(* Logix 5000 project; controller UOWHF Emulate 5570 rev 30.12; software revision 30.00 *) (continued)
   		UOWHF_Add_c.2:=UOWHF_Result[2].31;
   		UOWHF_Result[2].31:=0;
   		UOWHF_Result[3]:=UOWHF_Result[3] + 1798644847+UOWHF_Add_c;
   		UOWHF_Add_c.3:=UOWHF_Result[3].31;
   		UOWHF_Result[3].31:=0;
   		UOWHF_Result[4]:=UOWHF_Result[4] + 304175449+UOWHF_Add_c;
   		UOWHF_Add_c.4:=UOWHF_Result[4].31;
   		UOWHF_Result[4].31:=0;
   	End_If;
   	If UOWHF_Msg[2].[30] Then
   		UOWHF_Result[0]:=UOWHF_Result[0] + 1161935431+UOWHF_Add_c;
   		UOWHF_Add_c.0:=UOWHF_Result[0].31;
   		UOWHF_Result[0].31:=0;
   		UOWHF_Result[1]:=UOWHF_Result[1] + 944693816+UOWHF_Add_c;
   		UOWHF_Add_c.1:=UOWHF_Result[1].31;
   		UOWHF_Result[1].31:=0;
   		UOWHF_Result[2]:=UOWHF_Result[2] + 1100985340+UOWHF_Add_c;
   		UOWHF_Add_c.2:=UOWHF_Result[2].31;
   		UOWHF_Result[2].31:=0;
   		UOWHF_Result[3]:=UOWHF_Result[3] + 216963659+UOWHF_Add_c;
   		UOWHF_Add_c.3:=UOWHF_Result[3].31;
   		UOWHF_Result[3].31:=0;
   		UOWHF_Result[4]:=UOWHF_Result[4] + 89876541+UOWHF_Add_c;
   		UOWHF_Add_c.4:=UOWHF_Result[4].31;
   		UOWHF_Result[4].31:=0;
   	End_If;
   	If UOWHF_Msg[2].[31] Then
   		UOWHF_Result[0]:=UOWHF_Result[0] + 1158699558+UOWHF_Add_c;
   		UOWHF_Add_c.0:=UOWHF_Result[0].31;
   		UOWHF_Result[0].31:=0;
   		UOWHF_Result[1]:=UOWHF_Result[1] + 148835756+UOWHF_Add_c;
   		UOWHF_Add_c.1:=UOWHF_Result[1].31;
   		UOWHF_Result[1].31:=0;
   		UOWHF_Result[2]:=UOWHF_Result[2] + 32681667+UOWHF_Add_c;
   		UOWHF_Add_c.2:=UOWHF_Result[2].31;
   		UOWHF_Result[2].31:=0;
   		UOWHF_Result[3]:=UOWHF_Result[3] + 636137273+UOWHF_Add_c;
   		UOWHF_Add_c.3:=UOWHF_Result[3].31;
   		UOWHF_Result[3].31:=0;
   		UOWHF_Result[4]:=UOWHF_Result[4] + 1474642829+UOWHF_Add_c;
   		UOWHF_Add_c.4:=UOWHF_Result[4].31;
   		UOWHF_Result[4].31:=0;
   	End_If;
   	If UOWHF_Msg[3].[0] Then
   		UOWHF_Result[0]:=UOWHF_Result[0] + 1085349533+UOWHF_Add_c;
   		UOWHF_Add_c.0:=UOWHF_Result[0].31;
   		UOWHF_Result[0].31:=0;
   		UOWHF_Result[1]:=UOWHF_Result[1] + 1302835678+UOWHF_Add_c;
   		UOWHF_Add_c.1:=UOWHF_Result[1].31;
   		UOWHF_Result[1].31:=0;
   		UOWHF_Result[2]:=UOWHF_Result[2] + 681913251+UOWHF_Add_c;
   		UOWHF_Add_c.2:=UOWHF_Result[2].31;
   		UOWHF_Result[2].31:=0;
   		UOWHF_Result[3]:=UOWHF_Result[3] + 723730247+UOWHF_Add_c;
   		UOWHF_Add_c.3:=UOWHF_Result[3].31;
   		UOWHF_Result[3].31:=0;
   		UOWHF_Result[4]:=UOWHF_Result[4] + 7919506+UOWHF_Add_c;
   		UOWHF_Add_c.4:=UOWHF_Result[4].31;
   		UOWHF_Result[4].31:=0;
   	End_If;
   	If UOWHF_Msg[3].[1] Then
   		UOWHF_Result[0]:=UOWHF_Result[0] + 1136561897+UOWHF_Add_c;
   		UOWHF_Add_c.0:=UOWHF_Result[0].31;
   		UOWHF_Result[0].31:=0;
   		UOWHF_Result[1]:=UOWHF_Result[1] + 1822763236+UOWHF_Add_c;
   		UOWHF_Add_c.1:=UOWHF_Result[1].31;
   		UOWHF_Result[1].31:=0;
   		UOWHF_Result[2]:=UOWHF_Result[2] + 2116802572+UOWHF_Add_c;
   		UOWHF_Add_c.2:=UOWHF_Result[2].31;
   		UOWHF_Result[2].31:=0;
   		UOWHF_Result[3]:=UOWHF_Result[3] + 595130731+UOWHF_Add_c;
   		UOWHF_Add_c.3:=UOWHF_Result[3].31;
   		UOWHF_Result[3].31:=0;
   		UOWHF_Result[4]:=UOWHF_Result[4] + 1143215041+UOWHF_Add_c;
   		UOWHF_Add_c.4:=UOWHF_Result[4].31;
   		UOWHF_Result[4].31:=0;
   	End_If;
   	If UOWHF_Msg[3].[2] Then
   		UOWHF_Result[0]:=UOWHF_Result[0] + 44711483+UOWHF_Add_c;
   		UOWHF_Add_c.0:=UOWHF_Result[0].31;
   		UOWHF_Result[0].31:=0;
   		UOWHF_Result[1]:=UOWHF_Result[1] + 757400375+UOWHF_Add_c;
   		UOWHF_Add_c.1:=UOWHF_Result[1].31;
   		UOWHF_Result[1].31:=0;
   		UOWHF_Result[2]:=UOWHF_Result[2] + 1986965253+UOWHF_Add_c;
   		UOWHF_Add_c.2:=UOWHF_Result[2].31;
   		UOWHF_Result[2].31:=0;
   		UOWHF_Result[3]:=UOWHF_Result[3] + 1261883823+UOWHF_Add_c;
   		UOWHF_Add_c.3:=UOWHF_Result[3].31;
   		UOWHF_Result[3].31:=0;
   		UOWHF_Result[4]:=UOWHF_Result[4] + 1629162798+UOWHF_Add_c;
   		UOWHF_Add_c.4:=UOWHF_Result[4].31;
   		UOWHF_Result[4].31:=0;
   	End_If;
   	If UOWHF_Msg[3].[3] Then
   		UOWHF_Result[0]:=UOWHF_Result[0] + 927773888+UOWHF_Add_c;
   		UOWHF_Add_c.0:=UOWHF_Result[0].31;
   		UOWHF_Result[0].31:=0;
   		UOWHF_Result[1]:=UOWHF_Result[1] + 406294431+UOWHF_Add_c;
   		UOWHF_Add_c.1:=UOWHF_Result[1].31;
   		UOWHF_Result[1].31:=0;
   		UOWHF_Result[2]:=UOWHF_Result[2] + 1401005734+UOWHF_Add_c;
   		UOWHF_Add_c.2:=UOWHF_Result[2].31;
   		UOWHF_Result[2].31:=0;
   		UOWHF_Result[3]:=UOWHF_Result[3] + 68199430+UOWHF_Add_c;
   		UOWHF_Add_c.3:=UOWHF_Result[3].31;
   		UOWHF_Result[3].31:=0;
   		UOWHF_Result[4]:=UOWHF_Result[4] + 19140251+UOWHF_Add_c;
   		UOWHF_Add_c.4:=UOWHF_Result[4].31;
   		UOWHF_Result[4].31:=0;
   	End_If;
   	If UOWHF_Msg[3].[4] Then
   		UOWHF_Result[0]:=UOWHF_Result[0] + 1465686449+UOWHF_Add_c;
   		UOWHF_Add_c.0:=UOWHF_Result[0].31;
   		UOWHF_Result[0].31:=0;
   		UOWHF_Result[1]:=UOWHF_Result[1] + 801325300+UOWHF_Add_c;
   		UOWHF_Add_c.1:=UOWHF_Result[1].31;
   		UOWHF_Result[1].31:=0;
   		UOWHF_Result[2]:=UOWHF_Result[2] + 1749934298+UOWHF_Add_c;
   		UOWHF_Add_c.2:=UOWHF_Result[2].31;
   		UOWHF_Result[2].31:=0;
   		UOWHF_Result[3]:=UOWHF_Result[3] + 134929849+UOWHF_Add_c;
   		UOWHF_Add_c.3:=UOWHF_Result[3].31;
   		UOWHF_Result[3].31:=0;
   		UOWHF_Result[4]:=UOWHF_Result[4] + 509005605+UOWHF_Add_c;
   		UOWHF_Add_c.4:=UOWHF_Result[4].31;
   		UOWHF_Result[4].31:=0;
   	End_If;
   	If UOWHF_Msg[3].[5] Then
   		UOWHF_Result[0]:=UOWHF_Result[0] + 1429827656+UOWHF_Add_c;
   		UOWHF_Add_c.0:=UOWHF_Result[0].31;
   		UOWHF_Result[0].31:=0;
   		UOWHF_Result[1]:=UOWHF_Result[1] + 1639863327+UOWHF_Add_c;
   		UOWHF_Add_c.1:=UOWHF_Result[1].31;
   		UOWHF_Result[1].31:=0;
   		UOWHF_Result[2]:=UOWHF_Result[2] + 934688503+UOWHF_Add_c;
   		UOWHF_Add_c.2:=UOWHF_Result[2].31;
   		UOWHF_Result[2].31:=0;
   		UOWHF_Result[3]:=UOWHF_Result[3] + 1162965313+UOWHF_Add_c;
   		UOWHF_Add_c.3:=UOWHF_Result[3].31;
   		UOWHF_Result[3].31:=0;
   		UOWHF_Result[4]:=UOWHF_Result[4] + 767744+UOWHF_Add_c;
   		UOWHF_Add_c.4:=UOWHF_Result[4].31;
   		UOWHF_Result[4].31:=0;
   	End_If;
   	If UOWHF_Msg[3].[6] Then
   		UOWHF_Result[0]:=UOWHF_Result[0] + 2104448245+UOWHF_Add_c;
   		UOWHF_Add_c.0:=UOWHF_Result[0].31;
   		UOWHF_Result[0].31:=0;
   		UOWHF_Result[1]:=UOWHF_Result[1] + 1893133446+UOWHF_Add_c;
   		UOWHF_Add_c.1:=UOWHF_Result[1].31;
   		UOWHF_Result[1].31:=0;
   		UOWHF_Result[2]:=UOWHF_Result[2] + 1965489067+UOWHF_Add_c;
   		UOWHF_Add_c.2:=UOWHF_Result[2].31;
   		UOWHF_Result[2].31:=0;
   		UOWHF_Result[3]:=UOWHF_Result[3] + 87146528+UOWHF_Add_c;
   		UOWHF_Add_c.3:=UOWHF_Result[3].31;
   		UOWHF_Result[3].31:=0;
   		UOWHF_Result[4]:=UOWHF_Result[4] + 373668245+UOWHF_Add_c;
   		UOWHF_Add_c.4:=UOWHF_Result[4].31;
   		UOWHF_Result[4].31:=0;
   	End_If;
   	If UOWHF_Msg[3].[7] Then
   		UOWHF_Result[0]:=UOWHF_Result[0] + 421829896+UOWHF_Add_c;
   		UOWHF_Add_c.0:=UOWHF_Result[0].31;
   		UOWHF_Result[0].31:=0;
   		UOWHF_Result[1]:=UOWHF_Result[1] + 1596327164+UOWHF_Add_c;
   		UOWHF_Add_c.1:=UOWHF_Result[1].31;
   		UOWHF_Result[1].31:=0;
   		UOWHF_Result[2]:=UOWHF_Result[2] + 1881340037+UOWHF_Add_c;
   		UOWHF_Add_c.2:=UOWHF_Result[2].31;
   		UOWHF_Result[2].31:=0;
   		UOWHF_Result[3]:=UOWHF_Result[3] + 605100392+UOWHF_Add_c;
   		UOWHF_Add_c.3:=UOWHF_Result[3].31;
   		UOWHF_Result[3].31:=0;
   		UOWHF_Result[4]:=UOWHF_Result[4] + 1262662835+UOWHF_Add_c;
   		UOWHF_Add_c.4:=UOWHF_Result[4].31;
   		UOWHF_Result[4].31:=0;
   	End_If;
   	If UOWHF_Msg[3].[8] Then
   		UOWHF_Result[0]:=UOWHF_Result[0] + 316065492+UOWHF_Add_c;
   		UOWHF_Add_c.0:=UOWHF_Result[0].31;
   		UOWHF_Result[0].31:=0;
   		UOWHF_Result[1]:=UOWHF_Result[1] + 1543311762+UOWHF_Add_c;
   		UOWHF_Add_c.1:=UOWHF_Result[1].31;
   		UOWHF_Result[1].31:=0;
   		UOWHF_Result[2]:=UOWHF_Result[2] + 2044228187+UOWHF_Add_c;
   		UOWHF_Add_c.2:=UOWHF_Result[2].31;
   		UOWHF_Result[2].31:=0;
   		UOWHF_Result[3]:=UOWHF_Result[3] + 1763648339+UOWHF_Add_c;
   		UOWHF_Add_c.3:=UOWHF_Result[3].31;
   		UOWHF_Result[3].31:=0;
   		UOWHF_Result[4]:=UOWHF_Result[4] + 1866883199+UOWHF_Add_c;
   		UOWHF_Add_c.4:=UOWHF_Result[4].31;
   		UOWHF_Result[4].31:=0;
   	End_If;
   	If UOWHF_Msg[3].[9] Then
   		UOWHF_Result[0]:=UOWHF_Result[0] + 1787911426+UOWHF_Add_c;
   		UOWHF_Add_c.0:=UOWHF_Result[0].31;
   		UOWHF_Result[0].31:=0;
   		UOWHF_Result[1]:=UOWHF_Result[1] + 234471005+UOWHF_Add_c;
   		UOWHF_Add_c.1:=UOWHF_Result[1].31;
   		UOWHF_Result[1].31:=0;
   		UOWHF_Result[2]:=UOWHF_Result[2] + 862019270+UOWHF_Add_c;
   		UOWHF_Add_c.2:=UOWHF_Result[2].31;
   		UOWHF_Result[2].31:=0;
   		UOWHF_Result[3]:=UOWHF_Result[3] + 134091934+UOWHF_Add_c;
   		UOWHF_Add_c.3:=UOWHF_Result[3].31;
   		UOWHF_Result[3].31:=0;
   		UOWHF_Result[4]:=UOWHF_Result[4] + 173621469+UOWHF_Add_c;
   		UOWHF_Add_c.4:=UOWHF_Result[4].31;
   		UOWHF_Result[4].31:=0;
   	End_If;
   	If UOWHF_Msg[3].[10] Then
   		UOWHF_Result[0]:=UOWHF_Result[0] + 271983001+UOWHF_Add_c;
   		UOWHF_Add_c.0:=UOWHF_Result[0].31;
   		UOWHF_Result[0].31:=0;
   		UOWHF_Result[1]:=UOWHF_Result[1] + 675410965+UOWHF_Add_c;
   		UOWHF_Add_c.1:=UOWHF_Result[1].31;
   		UOWHF_Result[1].31:=0;
   		UOWHF_Result[2]:=UOWHF_Result[2] + 2075099455+UOWHF_Add_c;
   		UOWHF_Add_c.2:=UOWHF_Result[2].31;
   		UOWHF_Result[2].31:=0;
   		UOWHF_Result[3]:=UOWHF_Result[3] + 755811265+UOWHF_Add_c;
   		UOWHF_Add_c.3:=UOWHF_Result[3].31;
   		UOWHF_Result[3].31:=0;
   		UOWHF_Result[4]:=UOWHF_Result[4] + 981610100+UOWHF_Add_c;
   		UOWHF_Add_c.4:=UOWHF_Result[4].31;
   		UOWHF_Result[4].31:=0;
   	End_If;
   	If UOWHF_Msg[3].[11] Then
   		UOWHF_Result[0]:=UOWHF_Result[0] + 2007459693+UOWHF_Add_c;
   		UOWHF_Add_c.0:=UOWHF_Result[0].31;
   		UOWHF_Result[0].31:=0;
   		UOWHF_Result[1]:=UOWHF_Result[1] + 1986772819+UOWHF_Add_c;
   		UOWHF_Add_c.1:=UOWHF_Result[1].31;
   		UOWHF_Result[1].31:=0;
   		UOWHF_Result[2]:=UOWHF_Result[2] + 529209603+UOWHF_Add_c;
   		UOWHF_Add_c.2:=UOWHF_Result[2].31;
   		UOWHF_Result[2].31:=0;
   		UOWHF_Result[3]:=UOWHF_Result[3] + 1850463358+UOWHF_Add_c;
   		UOWHF_Add_c.3:=UOWHF_Result[3].31;
   		UOWHF_Result[3].31:=0;
   		UOWHF_Result[4]:=UOWHF_Result[4] + 58342983+UOWHF_Add_c;
   		UOWHF_Add_c.4:=UOWHF_Result[4].31;
   		UOWHF_Result[4].31:=0;
   	End_If;
   	If UOWHF_Msg[3].[12] Then
   		UOWHF_Result[0]:=UOWHF_Result[0] + 1749062231+UOWHF_Add_c;
   		UOWHF_Add_c.0:=UOWHF_Result[0].31;
   		UOWHF_Result[0].31:=0;
   		UOWHF_Result[1]:=UOWHF_Result[1] + 1646985135+UOWHF_Add_c;
   		UOWHF_Add_c.1:=UOWHF_Result[1].31;
   		UOWHF_Result[1].31:=0;
   		UOWHF_Result[2]:=UOWHF_Result[2] + 1387540803+UOWHF_Add_c;
   		UOWHF_Add_c.2:=UOWHF_Result[2].31;
   		UOWHF_Result[2].31:=0;
   		UOWHF_Result[3]:=UOWHF_Result[3] + 157665719+UOWHF_Add_c;
   		UOWHF_Add_c.3:=UOWHF_Result[3].31;
   		UOWHF_Result[3].31:=0;
   		UOWHF_Result[4]:=UOWHF_Result[4] + 458465077+UOWHF_Add_c;
   		UOWHF_Add_c.4:=UOWHF_Result[4].31;
   		UOWHF_Result[4].31:=0;
   	End_If;
   	If UOWHF_Msg[3].[13] Then
   		UOWHF_Result[0]:=UOWHF_Result[0] + 302675244+UOWHF_Add_c;
   		UOWHF_Add_c.0:=UOWHF_Result[0].31;
   		UOWHF_Result[0].31:=0;
   		UOWHF_Result[1]:=UOWHF_Result[1] + 1351639650+UOWHF_Add_c;
   		UOWHF_Add_c.1:=UOWHF_Result[1].31;
   		UOWHF_Result[1].31:=0;
   		UOWHF_Result[2]:=UOWHF_Result[2] + 930571861+UOWHF_Add_c;
   		UOWHF_Add_c.2:=UOWHF_Result[2].31;
   		UOWHF_Result[2].31:=0;
   		UOWHF_Result[3]:=UOWHF_Result[3] + 2102488550+UOWHF_Add_c;
   		UOWHF_Add_c.3:=UOWHF_Result[3].31;
   		UOWHF_Result[3].31:=0;
   		UOWHF_Result[4]:=UOWHF_Result[4] + 176477540+UOWHF_Add_c;
   		UOWHF_Add_c.4:=UOWHF_Result[4].31;
   		UOWHF_Result[4].31:=0;
   	End_If;
   	If UOWHF_Msg[3].[14] Then
   		UOWHF_Result[0]:=UOWHF_Result[0] + 286779437+UOWHF_Add_c;
   		UOWHF_Add_c.0:=UOWHF_Result[0].31;
   		UOWHF_Result[0].31:=0;
   		UOWHF_Result[1]:=UOWHF_Result[1] + 1779831145+UOWHF_Add_c;
   		UOWHF_Add_c.1:=UOWHF_Result[1].31;
   		UOWHF_Result[1].31:=0;
   		UOWHF_Result[2]:=UOWHF_Result[2] + 457655217+UOWHF_Add_c;
   		UOWHF_Add_c.2:=UOWHF_Result[2].31;
   		UOWHF_Result[2].31:=0;
   		UOWHF_Result[3]:=UOWHF_Result[3] + 1853803003+UOWHF_Add_c;
   		UOWHF_Add_c.3:=UOWHF_Result[3].31;
   		UOWHF_Result[3].31:=0;
   		UOWHF_Result[4]:=UOWHF_Result[4] + 1073511598+UOWHF_Add_c;
   		UOWHF_Add_c.4:=UOWHF_Result[4].31;
   		UOWHF_Result[4].31:=0;
   	End_If;
   	If UOWHF_Msg[3].[15] Then
   		UOWHF_Result[0]:=UOWHF_Result[0] + 1600464813+UOWHF_Add_c;
   		UOWHF_Add_c.0:=UOWHF_Result[0].31;
   		UOWHF_Result[0].31:=0;
   		UOWHF_Result[1]:=UOWHF_Result[1] + 415810416+UOWHF_Add_c;
   		UOWHF_Add_c.1:=UOWHF_Result[1].31;
   		UOWHF_Result[1].31:=0;
   		UOWHF_Result[2]:=UOWHF_Result[2] + 1110267176+UOWHF_Add_c;
   		UOWHF_Add_c.2:=UOWHF_Result[2].31;
   		UOWHF_Result[2].31:=0;
   		UOWHF_Result[3]:=UOWHF_Result[3] + 681690366+UOWHF_Add_c;
   		UOWHF_Add_c.3:=UOWHF_Result[3].31;
   		UOWHF_Result[3].31:=0;
   		UOWHF_Result[4]:=UOWHF_Result[4] + 89351772+UOWHF_Add_c;
   		UOWHF_Add_c.4:=UOWHF_Result[4].31;
   		UOWHF_Result[4].31:=0;
   	End_If;
   	If UOWHF_Msg[3].[16] Then
   		UOWHF_Result[0]:=UOWHF_Result[0] + 1422191011+UOWHF_Add_c;
   		UOWHF_Add_c.0:=UOWHF_Result[0].31;
   		UOWHF_Result[0].31:=0;
   		UOWHF_Result[1]:=UOWHF_Result[1] + 792068346+UOWHF_Add_c;
   		UOWHF_Add_c.1:=UOWHF_Result[1].31;
   		UOWHF_Result[1].31:=0;
   		UOWHF_Result[2]:=UOWHF_Result[2] + 931635063+UOWHF_Add_c;
   		UOWHF_Add_c.2:=UOWHF_Result[2].31;
   		UOWHF_Result[2].31:=0;
   		UOWHF_Result[3]:=UOWHF_Result[3] + 658957375+UOWHF_Add_c;
   		UOWHF_Add_c.3:=UOWHF_Result[3].31;
   		UOWHF_Result[3].31:=0;
   		UOWHF_Result[4]:=UOWHF_Result[4] + 1912632671+UOWHF_Add_c;
   		UOWHF_Add_c.4:=UOWHF_Result[4].31;
   		UOWHF_Result[4].31:=0;
   	End_If;
   	If UOWHF_Msg[3].[17] Then
   		UOWHF_Result[0]:=UOWHF_Result[0] + 1459819100+UOWHF_Add_c;
   		UOWHF_Add_c.0:=UOWHF_Result[0].31;
   		UOWHF_Result[0].31:=0;
   		UOWHF_Result[1]:=UOWHF_Result[1] + 444070721+UOWHF_Add_c;
   		UOWHF_Add_c.1:=UOWHF_Result[1].31;
   		UOWHF_Result[1].31:=0;
   		UOWHF_Result[2]:=UOWHF_Result[2] + 1552170238+UOWHF_Add_c;
   		UOWHF_Add_c.2:=UOWHF_Result[2].31;
   		UOWHF_Result[2].31:=0;
   		UOWHF_Result[3]:=UOWHF_Result[3] + 1379870988+UOWHF_Add_c;
   		UOWHF_Add_c.3:=UOWHF_Result[3].31;
   		UOWHF_Result[3].31:=0;
   		UOWHF_Result[4]:=UOWHF_Result[4] + 1241938678+UOWHF_Add_c;
   		UOWHF_Add_c.4:=UOWHF_Result[4].31;
   		UOWHF_Result[4].31:=0;
   	End_If;
   	If UOWHF_Msg[3].[18] Then
   		UOWHF_Result[0]:=UOWHF_Result[0] + 1537182853+UOWHF_Add_c;
   		UOWHF_Add_c.0:=UOWHF_Result[0].31;
   		UOWHF_Result[0].31:=0;
   		UOWHF_Result[1]:=UOWHF_Result[1] + 821913954+UOWHF_Add_c;
   		UOWHF_Add_c.1:=UOWHF_Result[1].31;
   		UOWHF_Result[1].31:=0;
   		UOWHF_Result[2]:=UOWHF_Result[2] + 2085504538+UOWHF_Add_c;
   		UOWHF_Add_c.2:=UOWHF_Result[2].31;
   		UOWHF_Result[2].31:=0;
   		UOWHF_Result[3]:=UOWHF_Result[3] + 349054710+UOWHF_Add_c;
   		UOWHF_Add_c.3:=UOWHF_Result[3].31;
   		UOWHF_Result[3].31:=0;
   		UOWHF_Result[4]:=UOWHF_Result[4] + 282436828+UOWHF_Add_c;
   		UOWHF_Add_c.4:=UOWHF_Result[4].31;
   		UOWHF_Result[4].31:=0;
   	End_If;
   	If UOWHF_Msg[3].[19] Then
   		UOWHF_Result[0]:=UOWHF_Result[0] + 190091110+UOWHF_Add_c;
   		UOWHF_Add_c.0:=UOWHF_Result[0].31;
   		UOWHF_Result[0].31:=0;
   		UOWHF_Result[1]:=UOWHF_Result[1] + 824558472+UOWHF_Add_c;
   		UOWHF_Add_c.1:=UOWHF_Result[1].31;
   		UOWHF_Result[1].31:=0;
   		UOWHF_Result[2]:=UOWHF_Result[2] + 165095409+UOWHF_Add_c;
   		UOWHF_Add_c.2:=UOWHF_Result[2].31;
   		UOWHF_Result[2].31:=0;
   		UOWHF_Result[3]:=UOWHF_Result[3] + 1237861916+UOWHF_Add_c;
   		UOWHF_Add_c.3:=UOWHF_Result[3].31;
   		UOWHF_Result[3].31:=0;
   		UOWHF_Result[4]:=UOWHF_Result[4] + 193118018+UOWHF_Add_c;
   		UOWHF_Add_c.4:=UOWHF_Result[4].31;
   		UOWHF_Result[4].31:=0;
   	End_If;
   	If UOWHF_Msg[3].[20] Then
   		UOWHF_Result[0]:=UOWHF_Result[0] + 12764661+UOWHF_Add_c;
   		UOWHF_Add_c.0:=UOWHF_Result[0].31;
   		UOWHF_Result[0].31:=0;
   		UOWHF_Result[1]:=UOWHF_Result[1] + 2140015145+UOWHF_Add_c;
   		UOWHF_Add_c.1:=UOWHF_Result[1].31;
   		UOWHF_Result[1].31:=0;
   		UOWHF_Result[2]:=UOWHF_Result[2] + 1002316216+UOWHF_Add_c;
   		UOWHF_Add_c.2:=UOWHF_Result[2].31;
   		UOWHF_Result[2].31:=0;
   		UOWHF_Result[3]:=UOWHF_Result[3] + 487193130+UOWHF_Add_c;
   		UOWHF_Add_c.3:=UOWHF_Result[3].31;
   		UOWHF_Result[3].31:=0;
   		UOWHF_Result[4]:=UOWHF_Result[4] + 1676712644+UOWHF_Add_c;
   		UOWHF_Add_c.4:=UOWHF_Result[4].31;
   		UOWHF_Result[4].31:=0;
   	End_If;
   	If UOWHF_Msg[3].[21] Then
   		UOWHF_Result[0]:=UOWHF_Result[0] + 1907563985+UOWHF_Add_c;
   		UOWHF_Add_c.0:=UOWHF_Result[0].31;
   		UOWHF_Result[0].31:=0;
   		UOWHF_Result[1]:=UOWHF_Result[1] + 969114504+UOWHF_Add_c;
   		UOWHF_Add_c.1:=UOWHF_Result[1].31;
   		UOWHF_Result[1].31:=0;
   		UOWHF_Result[2]:=UOWHF_Result[2] + 520479841+UOWHF_Add_c;
   		UOWHF_Add_c.2:=UOWHF_Result[2].31;
   		UOWHF_Result[2].31:=0;
   		UOWHF_Result[3]:=UOWHF_Result[3] + 1257632595+UOWHF_Add_c;
   		UOWHF_Add_c.3:=UOWHF_Result[3].31;
   		UOWHF_Result[3].31:=0;
   		UOWHF_Result[4]:=UOWHF_Result[4] + 2109351775+UOWHF_Add_c;
   		UOWHF_Add_c.4:=UOWHF_Result[4].31;
   		UOWHF_Result[4].31:=0;
   	End_If;
   	If UOWHF_Msg[3].[22] Then
   		UOWHF_Result[0]:=UOWHF_Result[0] + 1053437027+UOWHF_Add_c;
   		UOWHF_Add_c.0:=UOWHF_Result[0].31;
   		UOWHF_Result[0].31:=0;
   		UOWHF_Result[1]:=UOWHF_Result[1] + 1848473161+UOWHF_Add_c;
   		UOWHF_Add_c.1:=UOWHF_Result[1].31;
   		UOWHF_Result[1].31:=0;
   		UOWHF_Result[2]:=UOWHF_Result[2] + 436614652+UOWHF_Add_c;
   		UOWHF_Add_c.2:=UOWHF_Result[2].31;
   		UOWHF_Result[2].31:=0;
   		UOWHF_Result[3]:=UOWHF_Result[3] + 141740774+UOWHF_Add_c;
   		UOWHF_Add_c.3:=UOWHF_Result[3].31;
   		UOWHF_Result[3].31:=0;
   		UOWHF_Result[4]:=UOWHF_Result[4] + 1110639400+UOWHF_Add_c;
   		UOWHF_Add_c.4:=UOWHF_Result[4].31;
   		UOWHF_Result[4].31:=0;
   	End_If;
   	If UOWHF_Msg[3].[23] Then
   		UOWHF_Result[0]:=UOWHF_Result[0] + 1424986516+UOWHF_Add_c;
   		UOWHF_Add_c.0:=UOWHF_Result[0].31;
   		UOWHF_Result[0].31:=0;
   		UOWHF_Result[1]:=UOWHF_Result[1] + 1637174944+UOWHF_Add_c;
   		UOWHF_Add_c.1:=UOWHF_Result[1].31;
   		UOWHF_Result[1].31:=0;
   		UOWHF_Result[2]:=UOWHF_Result[2] + 1728901188+UOWHF_Add_c;
   		UOWHF_Add_c.2:=UOWHF_Result[2].31;
   		UOWHF_Result[2].31:=0;
   		UOWHF_Result[3]:=UOWHF_Result[3] + 2136059085+UOWHF_Add_c;
   		UOWHF_Add_c.3:=UOWHF_Result[3].31;
   		UOWHF_Result[3].31:=0;
   		UOWHF_Result[4]:=UOWHF_Result[4] + 1296242343+UOWHF_Add_c;
   		UOWHF_Add_c.4:=UOWHF_Result[4].31;
   		UOWHF_Result[4].31:=0;
   	End_If;
   	If UOWHF_Msg[3].[24] Then
   		UOWHF_Result[0]:=UOWHF_Result[0] + 642610093+UOWHF_Add_c;
   		UOWHF_Add_c.0:=UOWHF_Result[0].31;
   		UOWHF_Result[0].31:=0;
   		UOWHF_Result[1]:=UOWHF_Result[1] + 352682737+UOWHF_Add_c;
   		UOWHF_Add_c.1:=UOWHF_Result[1].31;
   		UOWHF_Result[1].31:=0;
   		UOWHF_Result[2]:=UOWHF_Result[2] + 520559218+UOWHF_Add_c;
   		UOWHF_Add_c.2:=UOWHF_Result[2].31;
   		UOWHF_Result[2].31:=0;
   		UOWHF_Result[3]:=UOWHF_Result[3] + 860332796+UOWHF_Add_c;
   		UOWHF_Add_c.3:=UOWHF_Result[3].31;
   		UOWHF_Result[3].31:=0;
   		UOWHF_Result[4]:=UOWHF_Result[4] + 2130999817+UOWHF_Add_c;
   		UOWHF_Add_c.4:=UOWHF_Result[4].31;
   		UOWHF_Result[4].31:=0;
   	End_If;
   	If UOWHF_Msg[3].[25] Then
   		UOWHF_Result[0]:=UOWHF_Result[0] + 400835722+UOWHF_Add_c;
   		UOWHF_Add_c.0:=UOWHF_Result[0].31;
   		UOWHF_Result[0].31:=0;
   		UOWHF_Result[1]:=UOWHF_Result[1] + 94325367+UOWHF_Add_c;
   		UOWHF_Add_c.1:=UOWHF_Result[1].31;
   		UOWHF_Result[1].31:=0;
   		UOWHF_Result[2]:=UOWHF_Result[2] + 1951698740+UOWHF_Add_c;
   		UOWHF_Add_c.2:=UOWHF_Result[2].31;
   		UOWHF_Result[2].31:=0;
   		UOWHF_Result[3]:=UOWHF_Result[3] + 913446042+UOWHF_Add_c;
   		UOWHF_Add_c.3:=UOWHF_Result[3].31;
   		UOWHF_Result[3].31:=0;
   		UOWHF_Result[4]:=UOWHF_Result[4] + 465750883+UOWHF_Add_c;
   		UOWHF_Add_c.4:=UOWHF_Result[4].31;
   		UOWHF_Result[4].31:=0;
   	End_If;
   	If UOWHF_Msg[3].[26] Then
   		UOWHF_Result[0]:=UOWHF_Result[0] + 550639475+UOWHF_Add_c;
   		UOWHF_Add_c.0:=UOWHF_Result[0].31;
   		UOWHF_Result[0].31:=0;
   		UOWHF_Result[1]:=UOWHF_Result[1] + 766311515+UOWHF_Add_c;
   		UOWHF_Add_c.1:=UOWHF_Result[1].31;
   		UOWHF_Result[1].31:=0;
   		UOWHF_Result[2]:=UOWHF_Result[2] + 201914688+UOWHF_Add_c;
   		UOWHF_Add_c.2:=UOWHF_Result[2].31;
   		UOWHF_Result[2].31:=0;
   		UOWHF_Result[3]:=UOWHF_Result[3] + 1072080534+UOWHF_Add_c;
   		UOWHF_Add_c.3:=UOWHF_Result[3].31;
   		UOWHF_Result[3].31:=0;
   		UOWHF_Result[4]:=UOWHF_Result[4] + 539028112+UOWHF_Add_c;
   		UOWHF_Add_c.4:=UOWHF_Result[4].31;
   		UOWHF_Result[4].31:=0;
   	End_If;
   	If UOWHF_Msg[3].[27] Then
   		UOWHF_Result[0]:=UOWHF_Result[0] + 730868366+UOWHF_Add_c;
   		UOWHF_Add_c.0:=UOWHF_Result[0].31;
   		UOWHF_Result[0].31:=0;
   		UOWHF_Result[1]:=UOWHF_Result[1] + 1489762528+UOWHF_Add_c;
   		UOWHF_Add_c.1:=UOWHF_Result[1].31;
   		UOWHF_Result[1].31:=0;
   		UOWHF_Result[2]:=UOWHF_Result[2] + 115143668+UOWHF_Add_c;
   		UOWHF_Add_c.2:=UOWHF_Result[2].31;
   		UOWHF_Result[2].31:=0;
   		UOWHF_Result[3]:=UOWHF_Result[3] + 1979129004+UOWHF_Add_c;
   		UOWHF_Add_c.3:=UOWHF_Result[3].31;
   		UOWHF_Result[3].31:=0;
   		UOWHF_Result[4]:=UOWHF_Result[4] + 524515597+UOWHF_Add_c;
   		UOWHF_Add_c.4:=UOWHF_Result[4].31;
   		UOWHF_Result[4].31:=0;
   	End_If;
   	If UOWHF_Msg[3].[28] Then
   		UOWHF_Result[0]:=UOWHF_Result[0] + 422624123+UOWHF_Add_c;
   		UOWHF_Add_c.0:=UOWHF_Result[0].31;
   		UOWHF_Result[0].31:=0;
   		UOWHF_Result[1]:=UOWHF_Result[1] + 2085556493+UOWHF_Add_c;
   		UOWHF_Add_c.1:=UOWHF_Result[1].31;
   		UOWHF_Result[1].31:=0;
   		UOWHF_Result[2]:=UOWHF_Result[2] + 2061386247+UOWHF_Add_c;
   		UOWHF_Add_c.2:=UOWHF_Result[2].31;
   		UOWHF_Result[2].31:=0;
   		UOWHF_Result[3]:=UOWHF_Result[3] + 104622945+UOWHF_Add_c;
   		UOWHF_Add_c.3:=UOWHF_Result[3].31;
   		UOWHF_Result[3].31:=0;
   		UOWHF_Result[4]:=UOWHF_Result[4] + 1312719690+UOWHF_Add_c;
   		UOWHF_Add_c.4:=UOWHF_Result[4].31;
   		UOWHF_Result[4].31:=0;
   	End_If;
   	If UOWHF_Msg[3].[29] Then
   		UOWHF_Result[0]:=UOWHF_Result[0] + 1477103804+UOWHF_Add_c;
   		UOWHF_Add_c.0:=UOWHF_Result[0].31;
   		UOWHF_Result[0].31:=0;
   		UOWHF_Result[1]:=UOWHF_Result[1] + 1207034729+UOWHF_Add_c;
   		UOWHF_Add_c.1:=UOWHF_Result[1].31;
   		UOWHF_Result[1].31:=0;
   		UOWHF_Result[2]:=UOWHF_Result[2] + 125218042+UOWHF_Add_c;
   		UOWHF_Add_c.2:=UOWHF_Result[2].31;
   		UOWHF_Result[2].31:=0;
   		UOWHF_Result[3]:=UOWHF_Result[3] + 1252411627+UOWHF_Add_c;
   		UOWHF_Add_c.3:=UOWHF_Result[3].31;
   		UOWHF_Result[3].31:=0;
   		UOWHF_Result[4]:=UOWHF_Result[4] + 1395004731+UOWHF_Add_c;
   		UOWHF_Add_c.4:=UOWHF_Result[4].31;
   		UOWHF_Result[4].31:=0;
   	End_If;
   	If UOWHF_Msg[3].[30] Then
   		UOWHF_Result[0]:=UOWHF_Result[0] + 389079095+UOWHF_Add_c;
   		UOWHF_Add_c.0:=UOWHF_Result[0].31;
   		UOWHF_Result[0].31:=0;
   		UOWHF_Result[1]:=UOWHF_Result[1] + 898153102+UOWHF_Add_c;
   		UOWHF_Add_c.1:=UOWHF_Result[1].31;
   		UOWHF_Result[1].31:=0;
   		UOWHF_Result[2]:=UOWHF_Result[2] + 465664657+UOWHF_Add_c;
   		UOWHF_Add_c.2:=UOWHF_Result[2].31;
   		UOWHF_Result[2].31:=0;
   		UOWHF_Result[3]:=UOWHF_Result[3] + 1807585182+UOWHF_Add_c;
   		UOWHF_Add_c.3:=UOWHF_Result[3].31;
   		UOWHF_Result[3].31:=0;
   		UOWHF_Result[4]:=UOWHF_Result[4] + 1481633898+UOWHF_Add_c;
   		UOWHF_Add_c.4:=UOWHF_Result[4].31;
   		UOWHF_Result[4].31:=0;
   	End_If;
   	If UOWHF_Msg[3].[31] Then
   		UOWHF_Result[0]:=UOWHF_Result[0] + 483607650+UOWHF_Add_c;
   		UOWHF_Add_c.0:=UOWHF_Result[0].31;
   		UOWHF_Result[0].31:=0;
   		UOWHF_Result[1]:=UOWHF_Result[1] + 408888995+UOWHF_Add_c;
   		UOWHF_Add_c.1:=UOWHF_Result[1].31;
   		UOWHF_Result[1].31:=0;
   		UOWHF_Result[2]:=UOWHF_Result[2] + 1185305465+UOWHF_Add_c;
   		UOWHF_Add_c.2:=UOWHF_Result[2].31;
   		UOWHF_Result[2].31:=0;
   		UOWHF_Result[3]:=UOWHF_Result[3] + 169752186+UOWHF_Add_c;
   		UOWHF_Add_c.3:=UOWHF_Result[3].31;
   		UOWHF_Result[3].31:=0;
   		UOWHF_Result[4]:=UOWHF_Result[4] + 987073084+UOWHF_Add_c;
   		UOWHF_Add_c.4:=UOWHF_Result[4].31;
   		UOWHF_Result[4].31:=0;
   	End_If;
   	If UOWHF_Msg[4].[0] Then
   		UOWHF_Result[0]:=UOWHF_Result[0] + 1186018261+UOWHF_Add_c;
   		UOWHF_Add_c.0:=UOWHF_Result[0].31;
   		UOWHF_Result[0].31:=0;
   		UOWHF_Result[1]:=UOWHF_Result[1] + 1100688620+UOWHF_Add_c;
   		UOWHF_Add_c.1:=UOWHF_Result[1].31;
   		UOWHF_Result[1].31:=0;
   		UOWHF_Result[2]:=UOWHF_Result[2] + 1879258322+UOWHF_Add_c;
   		UOWHF_Add_c.2:=UOWHF_Result[2].31;
   		UOWHF_Result[2].31:=0;
   		UOWHF_Result[3]:=UOWHF_Result[3] + 771200367+UOWHF_Add_c;
   		UOWHF_Add_c.3:=UOWHF_Result[3].31;
   		UOWHF_Result[3].31:=0;
   		UOWHF_Result[4]:=UOWHF_Result[4] + 829145612+UOWHF_Add_c;
   		UOWHF_Add_c.4:=UOWHF_Result[4].31;
   		UOWHF_Result[4].31:=0;
   	End_If;
   	If UOWHF_Msg[4].[1] Then
   		UOWHF_Result[0]:=UOWHF_Result[0] + 1400433180+UOWHF_Add_c;
   		UOWHF_Add_c.0:=UOWHF_Result[0].31;
   		UOWHF_Result[0].31:=0;
   		UOWHF_Result[1]:=UOWHF_Result[1] + 2108209421+UOWHF_Add_c;
   		UOWHF_Add_c.1:=UOWHF_Result[1].31;
   		UOWHF_Result[1].31:=0;
   		UOWHF_Result[2]:=UOWHF_Result[2] + 946531010+UOWHF_Add_c;
   		UOWHF_Add_c.2:=UOWHF_Result[2].31;
   		UOWHF_Result[2].31:=0;
   		UOWHF_Result[3]:=UOWHF_Result[3] + 789709313+UOWHF_Add_c;
   		UOWHF_Add_c.3:=UOWHF_Result[3].31;
   		UOWHF_Result[3].31:=0;
   		UOWHF_Result[4]:=UOWHF_Result[4] + 298399889+UOWHF_Add_c;
   		UOWHF_Add_c.4:=UOWHF_Result[4].31;
   		UOWHF_Result[4].31:=0;
   	End_If;
   	If UOWHF_Msg[4].[2] Then
   		UOWHF_Result[0]:=UOWHF_Result[0] + 1193720141+UOWHF_Add_c;
   		UOWHF_Add_c.0:=UOWHF_Result[0].31;
   		UOWHF_Result[0].31:=0;
   		UOWHF_Result[1]:=UOWHF_Result[1] + 1274568895+UOWHF_Add_c;
   		UOWHF_Add_c.1:=UOWHF_Result[1].31;
   		UOWHF_Result[1].31:=0;
   		UOWHF_Result[2]:=UOWHF_Result[2] + 941441387+UOWHF_Add_c;
   		UOWHF_Add_c.2:=UOWHF_Result[2].31;
   		UOWHF_Result[2].31:=0;
   		UOWHF_Result[3]:=UOWHF_Result[3] + 743461627+UOWHF_Add_c;
   		UOWHF_Add_c.3:=UOWHF_Result[3].31;
   		UOWHF_Result[3].31:=0;
   		UOWHF_Result[4]:=UOWHF_Result[4] + 1604901691+UOWHF_Add_c;
   		UOWHF_Add_c.4:=UOWHF_Result[4].31;
   		UOWHF_Result[4].31:=0;
   	End_If;
   	If UOWHF_Msg[4].[3] Then
   		UOWHF_Result[0]:=UOWHF_Result[0] + 2104945846+UOWHF_Add_c;
   		UOWHF_Add_c.0:=UOWHF_Result[0].31;
   		UOWHF_Result[0].31:=0;
   		UOWHF_Result[1]:=UOWHF_Result[1] + 1617034836+UOWHF_Add_c;
   		UOWHF_Add_c.1:=UOWHF_Result[1].31;
   		UOWHF_Result[1].31:=0;
   		UOWHF_Result[2]:=UOWHF_Result[2] + 2093569769+UOWHF_Add_c;
   		UOWHF_Add_c.2:=UOWHF_Result[2].31;
   		UOWHF_Result[2].31:=0;
   		UOWHF_Result[3]:=UOWHF_Result[3] + 1080990755+UOWHF_Add_c;
   		UOWHF_Add_c.3:=UOWHF_Result[3].31;
   		UOWHF_Result[3].31:=0;
   		UOWHF_Result[4]:=UOWHF_Result[4] + 46488863+UOWHF_Add_c;
   		UOWHF_Add_c.4:=UOWHF_Result[4].31;
   		UOWHF_Result[4].31:=0;
   	End_If;
   	If UOWHF_Msg[4].[4] Then
   		UOWHF_Result[0]:=UOWHF_Result[0] + 1659675590+UOWHF_Add_c;
   		UOWHF_Add_c.0:=UOWHF_Result[0].31;
   		UOWHF_Result[0].31:=0;
   		UOWHF_Result[1]:=UOWHF_Result[1] + 1304797753+UOWHF_Add_c;
   		UOWHF_Add_c.1:=UOWHF_Result[1].31;
   		UOWHF_Result[1].31:=0;
   		UOWHF_Result[2]:=UOWHF_Result[2] + 836907414+UOWHF_Add_c;
   		UOWHF_Add_c.2:=UOWHF_Result[2].31;
   		UOWHF_Result[2].31:=0;
   		UOWHF_Result[3]:=UOWHF_Result[3] + 1887621218+UOWHF_Add_c;
   		UOWHF_Add_c.3:=UOWHF_Result[3].31;
   		UOWHF_Result[3].31:=0;
   		UOWHF_Result[4]:=UOWHF_Result[4] + 1508845977+UOWHF_Add_c;
   		UOWHF_Add_c.4:=UOWHF_Result[4].31;
   		UOWHF_Result[4].31:=0;
   	End_If;
   	If UOWHF_Msg[4].[5] Then
   		UOWHF_Result[0]:=UOWHF_Result[0] + 644187969+UOWHF_Add_c;
   		UOWHF_Add_c.0:=UOWHF_Result[0].31;
   		UOWHF_Result[0].31:=0;
   		UOWHF_Result[1]:=UOWHF_Result[1] + 680978661+UOWHF_Add_c;
   		UOWHF_Add_c.1:=UOWHF_Result[1].31;
   		UOWHF_Result[1].31:=0;
   		UOWHF_Result[2]:=UOWHF_Result[2] + 530286153+UOWHF_Add_c;
   		UOWHF_Add_c.2:=UOWHF_Result[2].31;
   		UOWHF_Result[2].31:=0;
   		UOWHF_Result[3]:=UOWHF_Result[3] + 1054302806+UOWHF_Add_c;
   		UOWHF_Add_c.3:=UOWHF_Result[3].31;
   		UOWHF_Result[3].31:=0;
   		UOWHF_Result[4]:=UOWHF_Result[4] + 1379455094+UOWHF_Add_c;
   		UOWHF_Add_c.4:=UOWHF_Result[4].31;
   		UOWHF_Result[4].31:=0;
   	End_If;
   	If UOWHF_Msg[4].[6] Then
   		UOWHF_Result[0]:=UOWHF_Result[0] + 1797006456+UOWHF_Add_c;
   		UOWHF_Add_c.0:=UOWHF_Result[0].31;
   		UOWHF_Result[0].31:=0;
   		UOWHF_Result[1]:=UOWHF_Result[1] + 1671641212+UOWHF_Add_c;
   		UOWHF_Add_c.1:=UOWHF_Result[1].31;
   		UOWHF_Result[1].31:=0;
   		UOWHF_Result[2]:=UOWHF_Result[2] + 1471479868+UOWHF_Add_c;
   		UOWHF_Add_c.2:=UOWHF_Result[2].31;
   		UOWHF_Result[2].31:=0;
   		UOWHF_Result[3]:=UOWHF_Result[3] + 1312631408+UOWHF_Add_c;
   		UOWHF_Add_c.3:=UOWHF_Result[3].31;
   		UOWHF_Result[3].31:=0;
   		UOWHF_Result[4]:=UOWHF_Result[4] + 1423663426+UOWHF_Add_c;
   		UOWHF_Add_c.4:=UOWHF_Result[4].31;
   		UOWHF_Result[4].31:=0;
   	End_If;
   	If UOWHF_Msg[4].[7] Then
   		UOWHF_Result[0]:=UOWHF_Result[0] + 609168526+UOWHF_Add_c;
   		UOWHF_Add_c.0:=UOWHF_Result[0].31;
   		UOWHF_Result[0].31:=0;
   		UOWHF_Result[1]:=UOWHF_Result[1] + 478903215+UOWHF_Add_c;
   		UOWHF_Add_c.1:=UOWHF_Result[1].31;
   		UOWHF_Result[1].31:=0;
   		UOWHF_Result[2]:=UOWHF_Result[2] + 2135853958+UOWHF_Add_c;
   		UOWHF_Add_c.2:=UOWHF_Result[2].31;
   		UOWHF_Result[2].31:=0;
   		UOWHF_Result[3]:=UOWHF_Result[3] + 1732375759+UOWHF_Add_c;
   		UOWHF_Add_c.3:=UOWHF_Result[3].31;
   		UOWHF_Result[3].31:=0;
   		UOWHF_Result[4]:=UOWHF_Result[4] + 115158473+UOWHF_Add_c;
   		UOWHF_Add_c.4:=UOWHF_Result[4].31;
   		UOWHF_Result[4].31:=0;
   	End_If;
   	If UOWHF_Msg[4].[8] Then
   		UOWHF_Result[0]:=UOWHF_Result[0] + 1989798588+UOWHF_Add_c;
   		UOWHF_Add_c.0:=UOWHF_Result[0].31;
   		UOWHF_Result[0].31:=0;
   		UOWHF_Result[1]:=UOWHF_Result[1] + 591703516+UOWHF_Add_c;
   		UOWHF_Add_c.1:=UOWHF_Result[1].31;
   		UOWHF_Result[1].31:=0;
   		UOWHF_Result[2]:=UOWHF_Result[2] + 1328366246+UOWHF_Add_c;
   		UOWHF_Add_c.2:=UOWHF_Result[2].31;
   		UOWHF_Result[2].31:=0;
   		UOWHF_Result[3]:=UOWHF_Result[3] + 1055479196+UOWHF_Add_c;
   		UOWHF_Add_c.3:=UOWHF_Result[3].31;
   		UOWHF_Result[3].31:=0;
   		UOWHF_Result[4]:=UOWHF_Result[4] + 1638831242+UOWHF_Add_c;
   		UOWHF_Add_c.4:=UOWHF_Result[4].31;
   		UOWHF_Result[4].31:=0;
   	End_If;
   	If UOWHF_Msg[4].[9] Then
   		UOWHF_Result[0]:=UOWHF_Result[0] + 622406376+UOWHF_Add_c;
   		UOWHF_Add_c.0:=UOWHF_Result[0].31;
   		UOWHF_Result[0].31:=0;
   		UOWHF_Result[1]:=UOWHF_Result[1] + 302456745+UOWHF_Add_c;
   		UOWHF_Add_c.1:=UOWHF_Result[1].31;
   		UOWHF_Result[1].31:=0;
   		UOWHF_Result[2]:=UOWHF_Result[2] + 1004502914+UOWHF_Add_c;
   		UOWHF_Add_c.2:=UOWHF_Result[2].31;
   		UOWHF_Result[2].31:=0;
   		UOWHF_Result[3]:=UOWHF_Result[3] + 1944958998+UOWHF_Add_c;
   		UOWHF_Add_c.3:=UOWHF_Result[3].31;
   		UOWHF_Result[3].31:=0;
   		UOWHF_Result[4]:=UOWHF_Result[4] + 1457990763+UOWHF_Add_c;
   		UOWHF_Add_c.4:=UOWHF_Result[4].31;
   		UOWHF_Result[4].31:=0;
   	End_If;
   	If UOWHF_Msg[4].[10] Then
   		UOWHF_Result[0]:=UOWHF_Result[0] + 1190952435+UOWHF_Add_c;
   		UOWHF_Add_c.0:=UOWHF_Result[0].31;
   		UOWHF_Result[0].31:=0;
   		UOWHF_Result[1]:=UOWHF_Result[1] + 906321176+UOWHF_Add_c;
   		UOWHF_Add_c.1:=UOWHF_Result[1].31;
   		UOWHF_Result[1].31:=0;
   		UOWHF_Result[2]:=UOWHF_Result[2] + 1114856499+UOWHF_Add_c;
   		UOWHF_Add_c.2:=UOWHF_Result[2].31;
   		UOWHF_Result[2].31:=0;
   		UOWHF_Result[3]:=UOWHF_Result[3] + 2109990137+UOWHF_Add_c;
   		UOWHF_Add_c.3:=UOWHF_Result[3].31;
   		UOWHF_Result[3].31:=0;
   		UOWHF_Result[4]:=UOWHF_Result[4] + 2127466898+UOWHF_Add_c;
   		UOWHF_Add_c.4:=UOWHF_Result[4].31;
   		UOWHF_Result[4].31:=0;
   	End_If;
   	If UOWHF_Msg[4].[11] Then
   		UOWHF_Result[0]:=UOWHF_Result[0] + 1094778735+UOWHF_Add_c;
   		UOWHF_Add_c.0:=UOWHF_Result[0].31;
   		UOWHF_Result[0].31:=0;
   		UOWHF_Result[1]:=UOWHF_Result[1] + 920886974+UOWHF_Add_c;
   		UOWHF_Add_c.1:=UOWHF_Result[1].31;
   		UOWHF_Result[1].31:=0;
   		UOWHF_Result[2]:=UOWHF_Result[2] + 1275226437+UOWHF_Add_c;
   		UOWHF_Add_c.2:=UOWHF_Result[2].31;
   		UOWHF_Result[2].31:=0;
   		UOWHF_Result[3]:=UOWHF_Result[3] + 82556508+UOWHF_Add_c;
   		UOWHF_Add_c.3:=UOWHF_Result[3].31;
   		UOWHF_Result[3].31:=0;
   		UOWHF_Result[4]:=UOWHF_Result[4] + 977078858+UOWHF_Add_c;
   		UOWHF_Add_c.4:=UOWHF_Result[4].31;
   		UOWHF_Result[4].31:=0;
   	End_If;
   	If UOWHF_Msg[4].[12] Then
   		UOWHF_Result[0]:=UOWHF_Result[0] + 593744688+UOWHF_Add_c;
   		UOWHF_Add_c.0:=UOWHF_Result[0].31;
   		UOWHF_Result[0].31:=0;
   		UOWHF_Result[1]:=UOWHF_Result[1] + 1169255414+UOWHF_Add_c;
   		UOWHF_Add_c.1:=UOWHF_Result[1].31;
   		UOWHF_Result[1].31:=0;
   		UOWHF_Result[2]:=UOWHF_Result[2] + 51716405+UOWHF_Add_c;
   		UOWHF_Add_c.2:=UOWHF_Result[2].31;
   		UOWHF_Result[2].31:=0;
   		UOWHF_Result[3]:=UOWHF_Result[3] + 1207915051+UOWHF_Add_c;
